// TIA Portal project "Plc_KTKDL" (V19) (continued)
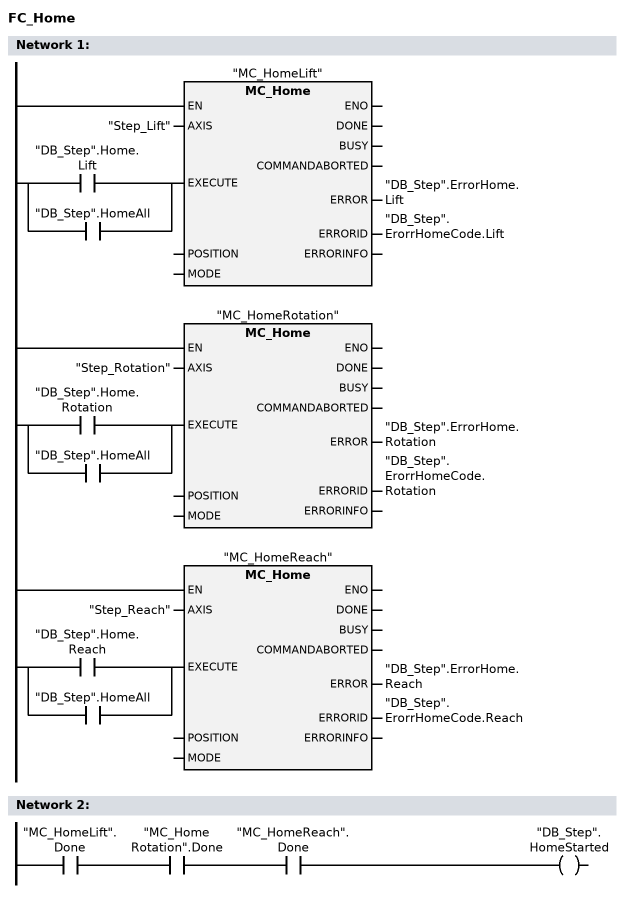
   "MC_HomeLift"(Axis := "Step_Lift",   // MC_Home
                 Execute := "DB_Step".Home.Lift OR "DB_Step".HomeAll,
                 Error => "DB_Step".ErrorHome.Lift,
                 ErrorID => "DB_Step".ErorrHomeCode.Lift);
   "MC_HomeRotation"(Axis := "Step_Rotation",   // MC_Home
                     Execute := "DB_Step".Home.Rotation OR "DB_Step".HomeAll,
                     Error => "DB_Step".ErrorHome.Rotation,
                     ErrorID => "DB_Step".ErorrHomeCode.Rotation);
   "MC_HomeReach"(Axis := "Step_Reach",   // MC_Home
                  Execute := "DB_Step".Home.Reach OR "DB_Step".HomeAll,
                  Error => "DB_Step".ErrorHome.Reach,
                  ErrorID => "DB_Step".ErorrHomeCode.Reach);
END_REGION

REGION Network 2
   RUNG wire#powerrail
      Contact( "MC_HomeLift".Done )
      Contact( "MC_HomeRotation".Done )
      Contact( "MC_HomeReach".Done )
      Coil( "DB_Step".HomeStarted )
   END_RUNG
   // the same network as SCL:
   "DB_Step".HomeStarted := "MC_HomeLift".Done AND "MC_HomeRotation".Done AND "MC_HomeReach".Done;
END_REGION
END_FUNCTION

FUNCTION "FC_Auto" : Void   // FC17, LAD
{ S7_Optimized_Access := 'TRUE' }
VERSION : 0.1
   VAR_TEMP   // added for the SCL form of the ladder/FBD networks
      _w1 : Bool;
      _w2 : Bool;
      _w3 : Bool;
      _w4 : Bool;
      _w5 : Bool;
      _w6 : Bool;
      _w7 : Bool;
      _w8 : Bool;
      _w9 : Bool;
      _w10 : Bool;
      _w11 : Bool;
      _w12 : Bool;
      _w13 : Bool;
      _w14 : Bool;
      _w15 : Bool;
      _w16 : Bool;
      _w17 : Bool;
      _w18 : Bool;
   END_VAR
BEGIN

REGION Network 1
   // 2 bước đầu là kiểm tra và set vận tốc
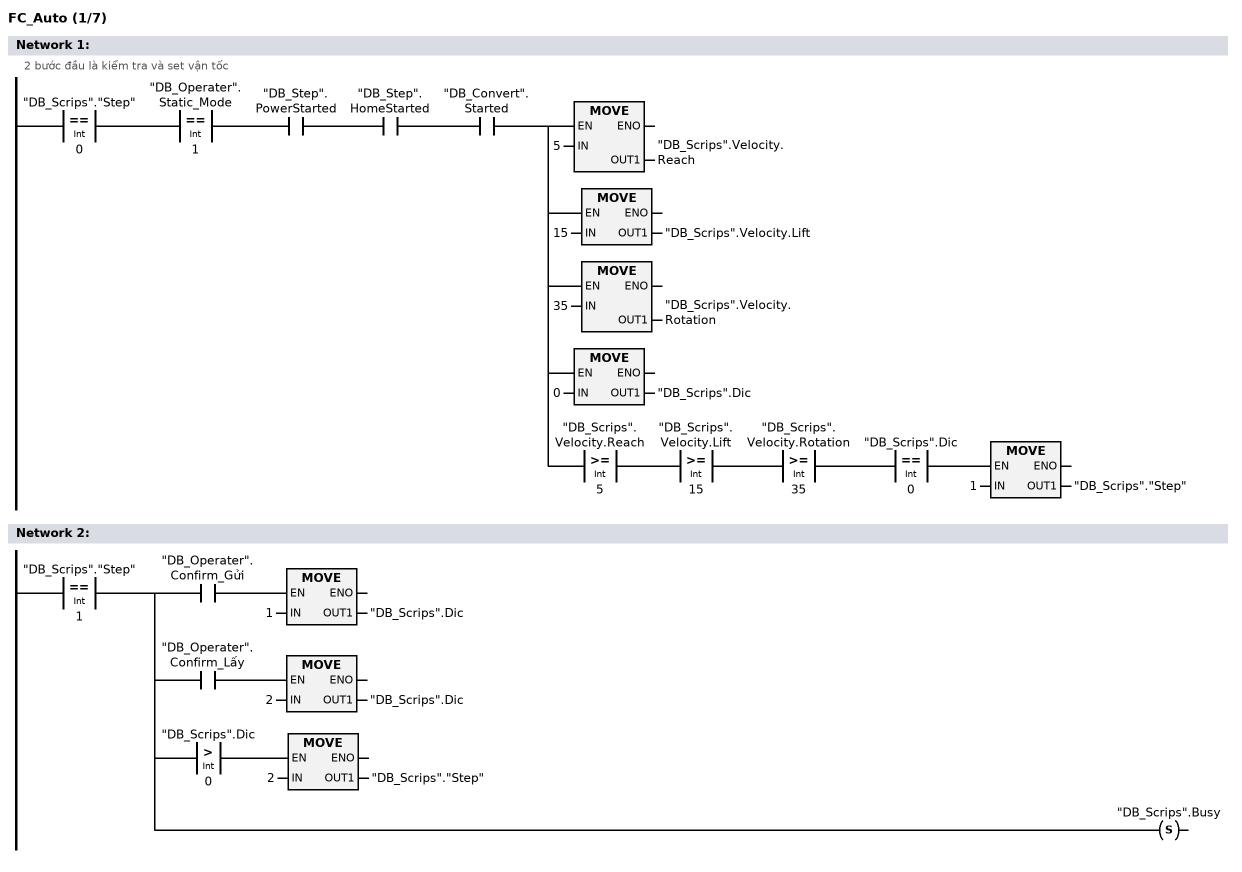
   RUNG wire#powerrail
      { S7_Templates := "SrcType := Int" } EQ_Contact(in1 := "DB_Scrips"."Step", in2 := 0)
      { S7_Templates := "SrcType := Int" } EQ_Contact(in1 := "DB_Operater".Static_Mode, in2 := 1)
      Contact( "DB_Step".PowerStarted )
      Contact( "DB_Step".HomeStarted )
      Contact( "DB_Convert".Started )
      wire#w1
      Move(in := 5, out1 => "DB_Scrips".Velocity.Reach)
   END_RUNG
   RUNG wire#w1
      Move(in := 15, out1 => "DB_Scrips".Velocity.Lift)
   END_RUNG
   RUNG wire#w1
      Move(in := 35, out1 => "DB_Scrips".Velocity.Rotation)
   END_RUNG
   RUNG wire#w1
      Move(in := 0, out1 => "DB_Scrips".Dic)
   END_RUNG
   RUNG wire#w1
      { S7_Templates := "SrcType := Int" } GE_Contact(in1 := "DB_Scrips".Velocity.Reach, in2 := 5)
      { S7_Templates := "SrcType := Int" } GE_Contact(in1 := "DB_Scrips".Velocity.Lift, in2 := 15)
      { S7_Templates := "SrcType := Int" } GE_Contact(in1 := "DB_Scrips".Velocity.Rotation, in2 := 35)
      { S7_Templates := "SrcType := Int" } EQ_Contact(in1 := "DB_Scrips".Dic, in2 := 0)
      Move(in := 1, out1 => "DB_Scrips"."Step")
   END_RUNG
   // the same network as SCL:
   #_w1 := ("DB_Scrips"."Step" = 0) AND ("DB_Operater".Static_Mode = 1) AND "DB_Step".PowerStarted AND "DB_Step".HomeStarted AND "DB_Convert".Started;
   IF #_w1 THEN
       "DB_Scrips".Velocity.Reach := 5;
       "DB_Scrips".Velocity.Lift := 15;
       "DB_Scrips".Velocity.Rotation := 35;
       "DB_Scrips".Dic := 0;
   END_IF;
   IF #_w1 AND ("DB_Scrips".Velocity.Reach >= 5) AND ("DB_Scrips".Velocity.Lift >= 15) AND ("DB_Scrips".Velocity.Rotation >= 35) AND ("DB_Scrips".Dic = 0) THEN
       "DB_Scrips"."Step" := 1;
   END_IF;
END_REGION

REGION Network 2
   RUNG wire#powerrail
      { S7_Templates := "SrcType := Int" } EQ_Contact(in1 := "DB_Scrips"."Step", in2 := 1)
      wire#w1
      Contact( "DB_Operater".Confirm_Gửi )
      Move(in := 1, out1 => "DB_Scrips".Dic)
   END_RUNG
   RUNG wire#w1
      Contact( "DB_Operater".Confirm_Lấy )
      Move(in := 2, out1 => "DB_Scrips".Dic)
   END_RUNG
   RUNG wire#w1
      { S7_Templates := "SrcType := Int" } GT_Contact(in1 := "DB_Scrips".Dic, in2 := 0)
      Move(in := 2, out1 => "DB_Scrips"."Step")
   END_RUNG
   RUNG wire#w1
      S_Coil( "DB_Scrips".Busy )
   END_RUNG
   // the same network as SCL:
   #_w1 := "DB_Scrips"."Step" = 1;
   IF #_w1 AND "DB_Operater".Confirm_Gửi THEN "DB_Scrips".Dic := 1; END_IF;
   IF #_w1 AND "DB_Operater".Confirm_Lấy THEN "DB_Scrips".Dic := 2; END_IF;
   IF #_w1 AND ("DB_Scrips".Dic > 0) THEN "DB_Scrips"."Step" := 2; END_IF;
   IF #_w1 THEN "DB_Scrips".Busy := TRUE; END_IF;
END_REGION

REGION Network 3
   // chưa làm logic lấy
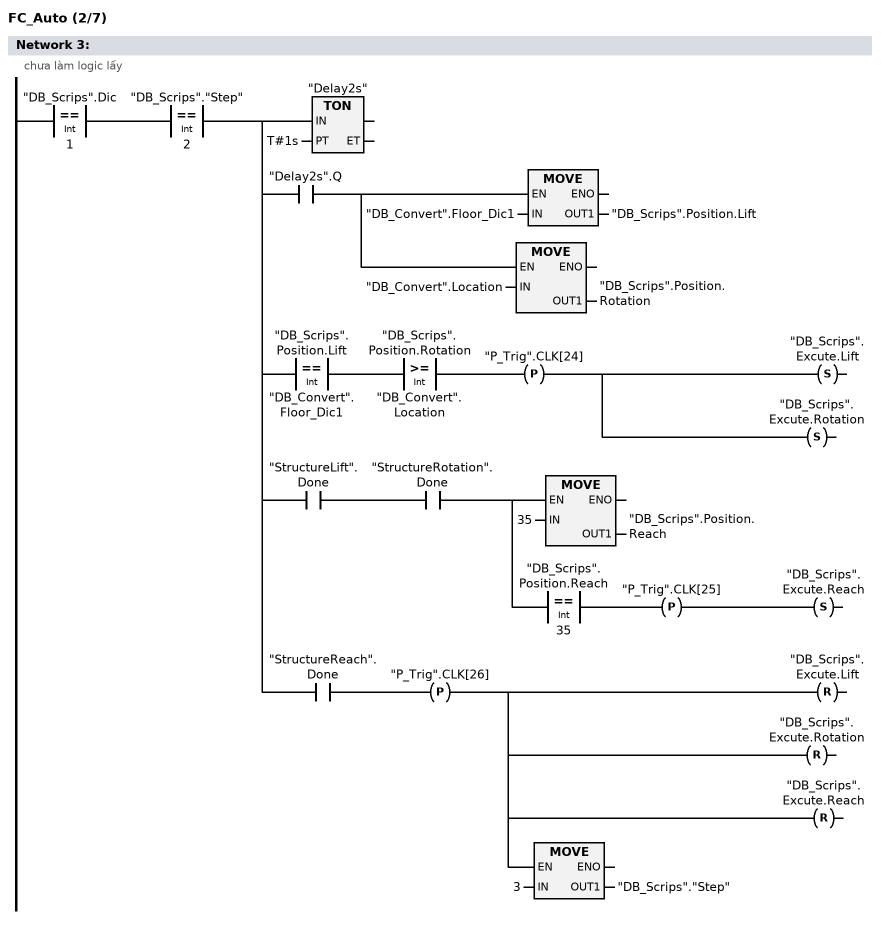
   #_w1 := ("DB_Scrips".Dic = 1) AND ("DB_Scrips"."Step" = 2);
   "Delay2s".TON(IN := #_w1, PT := T#1s);
   IF #_w1 AND "Delay2s".Q THEN
       "DB_Scrips".Position.Lift := "DB_Convert".Floor_Dic1;
       "DB_Scrips".Position.Rotation := "DB_Convert".Location;
   END_IF;
   #_w2 := #_w1 AND ("DB_Scrips".Position.Lift = "DB_Convert".Floor_Dic1) AND ("DB_Scrips".Position.Rotation >= "DB_Convert".Location);
   #_w3 := #_w2 AND NOT "P_Trig".CLK[24];   // rising edge
   "P_Trig".CLK[24] := #_w2;
   IF #_w3 THEN
       "DB_Scrips".Excute.Lift := TRUE;
       "DB_Scrips".Excute.Rotation := TRUE;
   END_IF;
   #_w4 := #_w1 AND "StructureLift".Done AND "StructureRotation".Done;
   IF #_w4 THEN "DB_Scrips".Position.Reach := 35; END_IF;
   #_w5 := #_w4 AND ("DB_Scrips".Position.Reach = 35);
   #_w6 := #_w5 AND NOT "P_Trig".CLK[25];   // rising edge
   "P_Trig".CLK[25] := #_w5;
   IF #_w6 THEN "DB_Scrips".Excute.Reach := TRUE; END_IF;
   #_w7 := #_w1 AND "StructureReach".Done;
   #_w8 := #_w7 AND NOT "P_Trig".CLK[26];   // rising edge
   "P_Trig".CLK[26] := #_w7;
   IF #_w8 THEN
       "DB_Scrips".Excute.Lift := FALSE;
       "DB_Scrips".Excute.Rotation := FALSE;
       "DB_Scrips".Excute.Reach := FALSE;
       "DB_Scrips"."Step" := 3;
   END_IF;
END_REGION

REGION Network 4
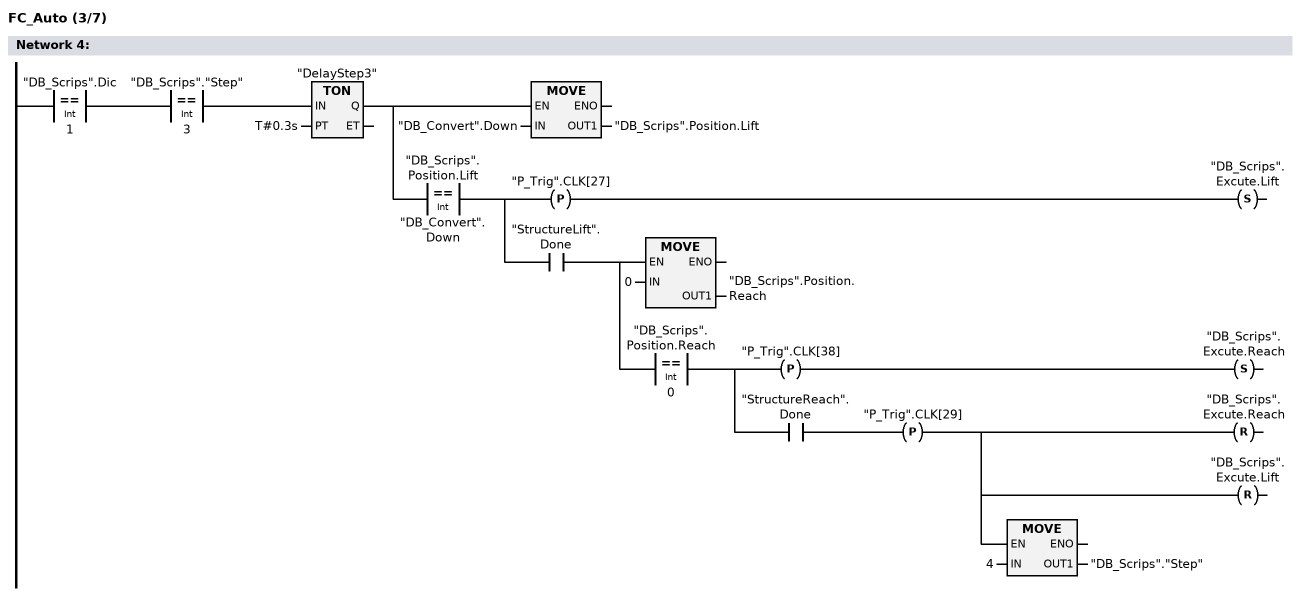
   "DelayStep3".TON(IN := ("DB_Scrips".Dic = 1) AND ("DB_Scrips"."Step" = 3), PT := T#0.3s);
   IF "DelayStep3".Q THEN "DB_Scrips".Position.Lift := "DB_Convert".Down; END_IF;
   #_w1 := "DelayStep3".Q AND ("DB_Scrips".Position.Lift = "DB_Convert".Down);
   #_w2 := #_w1 AND NOT "P_Trig".CLK[27];   // rising edge
   "P_Trig".CLK[27] := #_w1;
   IF #_w2 THEN "DB_Scrips".Excute.Lift := TRUE; END_IF;
   #_w3 := #_w1 AND "StructureLift".Done;
   IF #_w3 THEN "DB_Scrips".Position.Reach := 0; END_IF;
   #_w4 := #_w3 AND ("DB_Scrips".Position.Reach = 0);
   #_w5 := #_w4 AND NOT "P_Trig".CLK[38];   // rising edge
   "P_Trig".CLK[38] := #_w4;
   IF #_w5 THEN "DB_Scrips".Excute.Reach := TRUE; END_IF;
   #_w6 := #_w4 AND "StructureReach".Done;
   #_w7 := #_w6 AND NOT "P_Trig".CLK[29];   // rising edge
   "P_Trig".CLK[29] := #_w6;
   IF #_w7 THEN
       "DB_Scrips".Excute.Reach := FALSE;
       "DB_Scrips".Excute.Lift := FALSE;
       "DB_Scrips"."Step" := 4;
   END_IF;
END_REGION

REGION Network 5
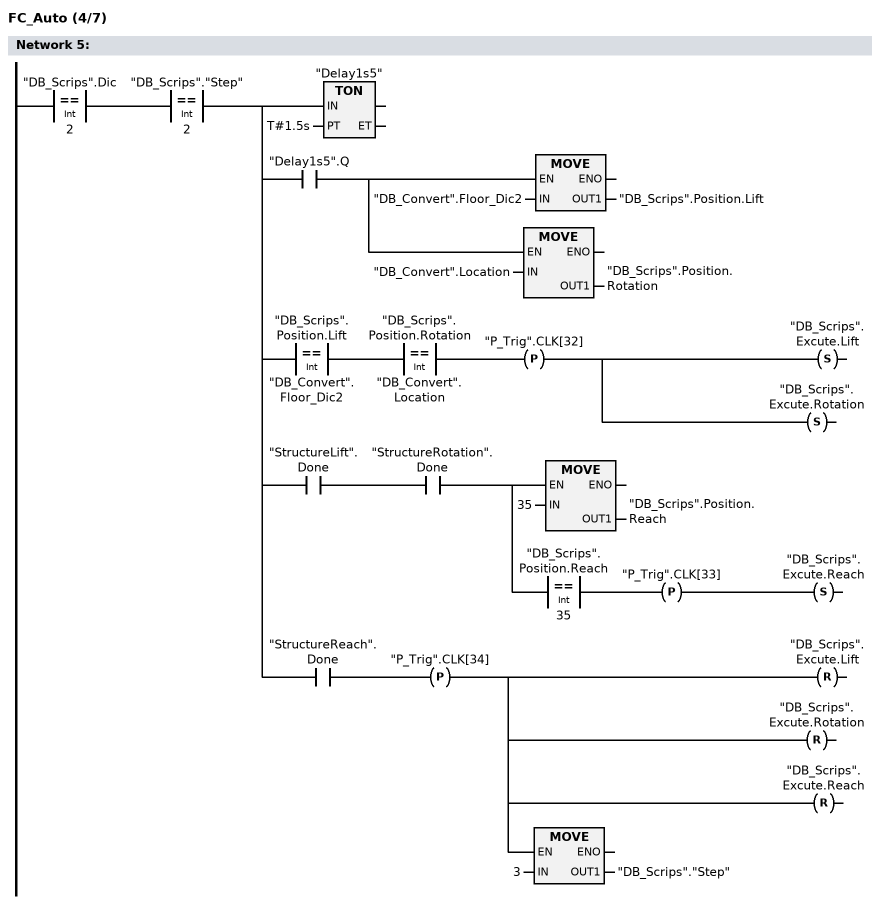
   #_w1 := ("DB_Scrips".Dic = 2) AND ("DB_Scrips"."Step" = 2);
   "Delay1s5".TON(IN := #_w1, PT := T#1.5s);
   IF #_w1 AND "Delay1s5".Q THEN
       "DB_Scrips".Position.Lift := "DB_Convert".Floor_Dic2;
       "DB_Scrips".Position.Rotation := "DB_Convert".Location;
   END_IF;
   #_w2 := #_w1 AND ("DB_Scrips".Position.Lift = "DB_Convert".Floor_Dic2) AND ("DB_Scrips".Position.Rotation = "DB_Convert".Location);
   #_w3 := #_w2 AND NOT "P_Trig".CLK[32];   // rising edge
   "P_Trig".CLK[32] := #_w2;
   IF #_w3 THEN
       "DB_Scrips".Excute.Lift := TRUE;
       "DB_Scrips".Excute.Rotation := TRUE;
   END_IF;
   #_w4 := #_w1 AND "StructureLift".Done AND "StructureRotation".Done;
   IF #_w4 THEN "DB_Scrips".Position.Reach := 35; END_IF;
   #_w5 := #_w4 AND ("DB_Scrips".Position.Reach = 35);
   #_w6 := #_w5 AND NOT "P_Trig".CLK[33];   // rising edge
   "P_Trig".CLK[33] := #_w5;
   IF #_w6 THEN "DB_Scrips".Excute.Reach := TRUE; END_IF;
   #_w7 := #_w1 AND "StructureReach".Done;
   #_w8 := #_w7 AND NOT "P_Trig".CLK[34];   // rising edge
   "P_Trig".CLK[34] := #_w7;
   IF #_w8 THEN
       "DB_Scrips".Excute.Lift := FALSE;
       "DB_Scrips".Excute.Rotation := FALSE;
       "DB_Scrips".Excute.Reach := FALSE;
       "DB_Scrips"."Step" := 3;
   END_IF;
END_REGION

REGION Network 6
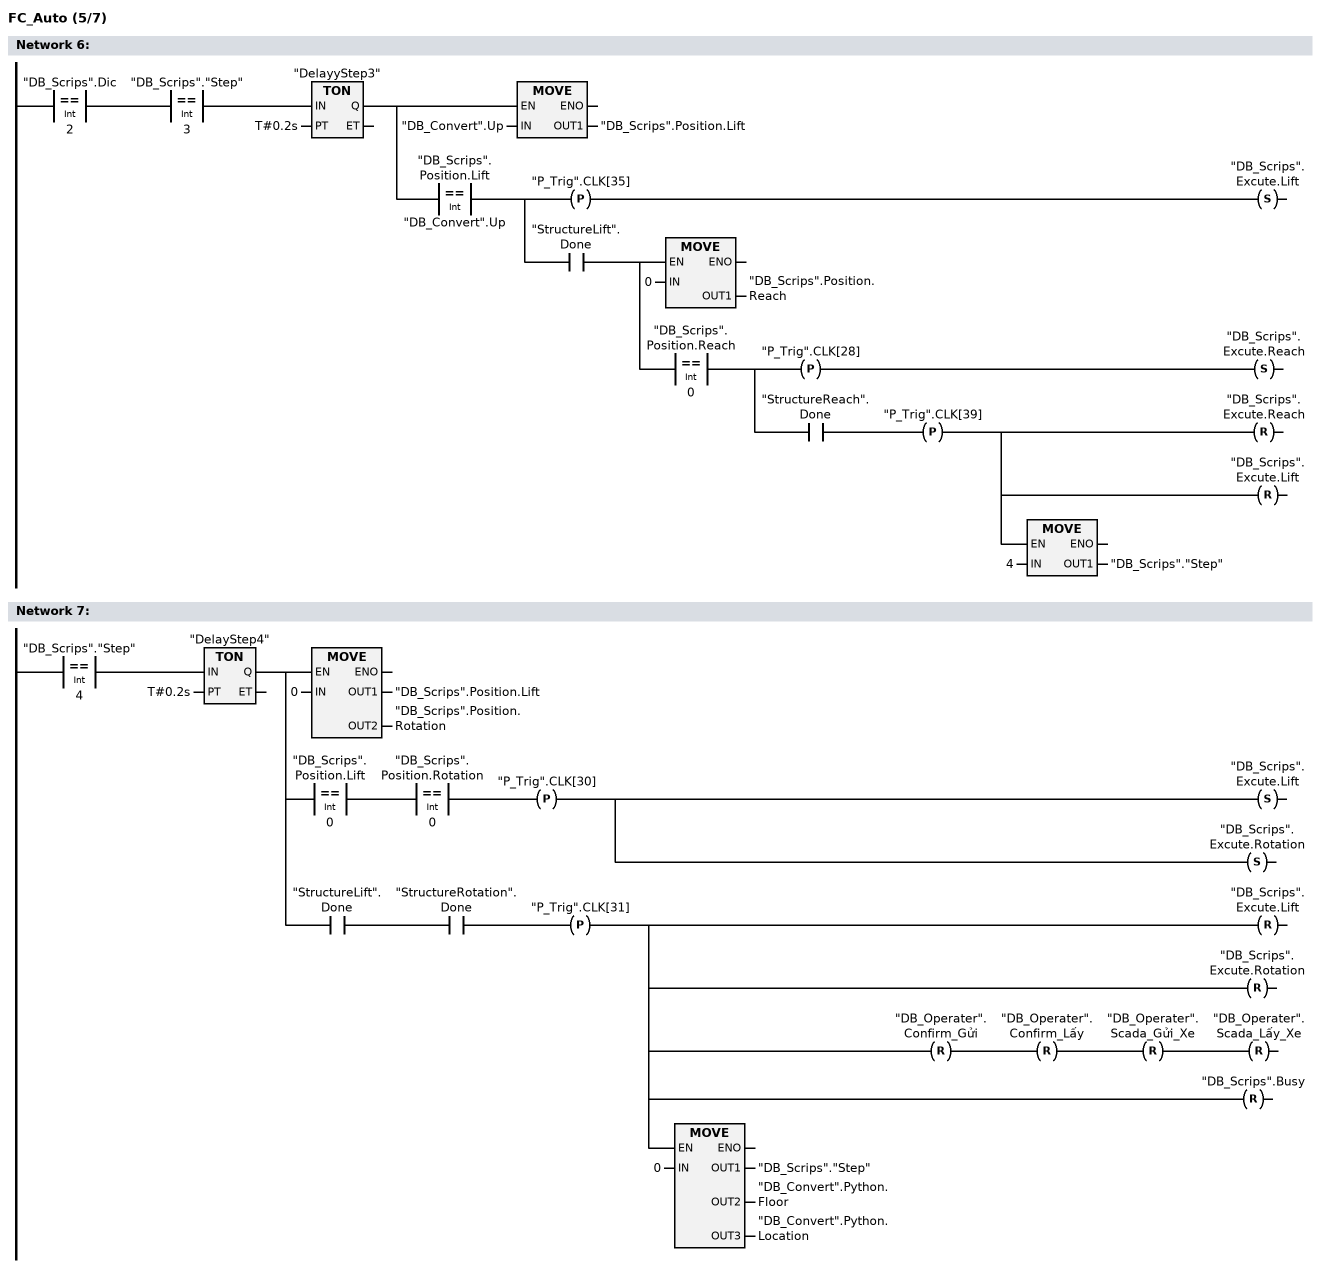
   "DelayyStep3".TON(IN := ("DB_Scrips".Dic = 2) AND ("DB_Scrips"."Step" = 3), PT := T#0.2s);
   IF "DelayyStep3".Q THEN "DB_Scrips".Position.Lift := "DB_Convert".Up; END_IF;
   #_w1 := "DelayyStep3".Q AND ("DB_Scrips".Position.Lift = "DB_Convert".Up);
   #_w2 := #_w1 AND NOT "P_Trig".CLK[35];   // rising edge
   "P_Trig".CLK[35] := #_w1;
   IF #_w2 THEN "DB_Scrips".Excute.Lift := TRUE; END_IF;
   #_w3 := #_w1 AND "StructureLift".Done;
   IF #_w3 THEN "DB_Scrips".Position.Reach := 0; END_IF;
   #_w4 := #_w3 AND ("DB_Scrips".Position.Reach = 0);
   #_w5 := #_w4 AND NOT "P_Trig".CLK[28];   // rising edge
   "P_Trig".CLK[28] := #_w4;
   IF #_w5 THEN "DB_Scrips".Excute.Reach := TRUE; END_IF;
   #_w6 := #_w4 AND "StructureReach".Done;
   #_w7 := #_w6 AND NOT "P_Trig".CLK[39];   // rising edge
   "P_Trig".CLK[39] := #_w6;
   IF #_w7 THEN
       "DB_Scrips".Excute.Reach := FALSE;
       "DB_Scrips".Excute.Lift := FALSE;
       "DB_Scrips"."Step" := 4;
   END_IF;
END_REGION

REGION Network 7
   "DelayStep4".TON(IN := "DB_Scrips"."Step" = 4, PT := T#0.2s);
   IF "DelayStep4".Q THEN
       "DB_Scrips".Position.Lift := 0;
       "DB_Scrips".Position.Rotation := 0;
   END_IF;
   #_w1 := "DelayStep4".Q AND ("DB_Scrips".Position.Lift = 0) AND ("DB_Scrips".Position.Rotation = 0);
   #_w2 := #_w1 AND NOT "P_Trig".CLK[30];   // rising edge
   "P_Trig".CLK[30] := #_w1;
   IF #_w2 THEN
       "DB_Scrips".Excute.Lift := TRUE;
       "DB_Scrips".Excute.Rotation := TRUE;
   END_IF;
   #_w3 := "DelayStep4".Q AND "StructureLift".Done AND "StructureRotation".Done;
   #_w4 := #_w3 AND NOT "P_Trig".CLK[31];   // rising edge
   "P_Trig".CLK[31] := #_w3;
   IF #_w4 THEN
       "DB_Scrips".Excute.Lift := FALSE;
       "DB_Scrips".Excute.Rotation := FALSE;
       "DB_Operater".Confirm_Gửi := FALSE;
       "DB_Operater".Confirm_Lấy := FALSE;
       "DB_Operater".Scada_Gửi_Xe := FALSE;
       "DB_Operater".Scada_Lấy_Xe := FALSE;
       "DB_Scrips".Busy := FALSE;
       "DB_Scrips"."Step" := 0;
       "DB_Convert".Python.Floor := 0;
       "DB_Convert".Python.Location := 0;
   END_IF;
END_REGION

REGION Network 9
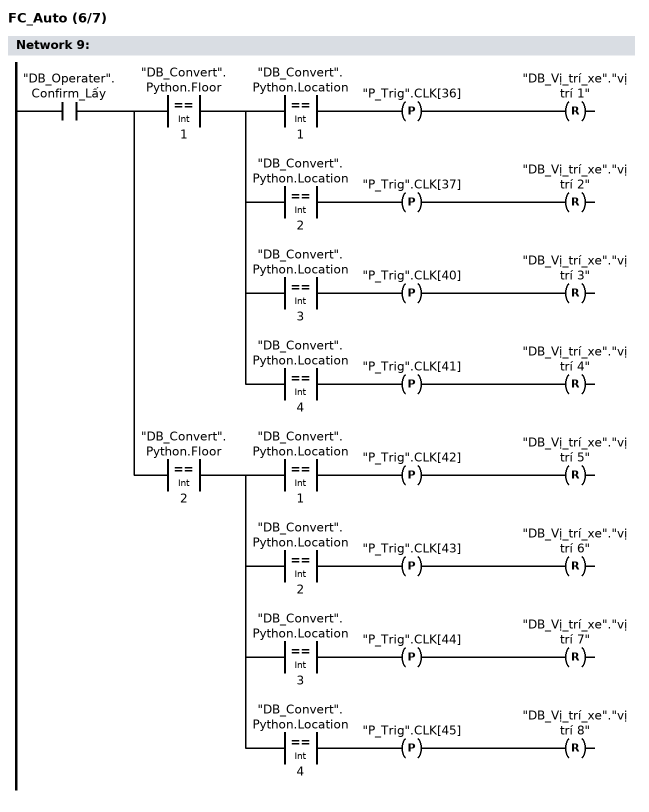
   RUNG wire#powerrail
      Contact( "DB_Operater".Confirm_Lấy )
      wire#w1
      { S7_Templates := "SrcType := Int" } EQ_Contact(in1 := "DB_Convert".Python.Floor, in2 := 1)
      wire#w2
      { S7_Templates := "SrcType := Int" } EQ_Contact(in1 := "DB_Convert".Python.Location, in2 := 1)
      P_Trig( "P_Trig".CLK[36] )
      R_Coil( "DB_Vị_trí_xe"."vị trí 1" )
   END_RUNG
   RUNG wire#w2
      { S7_Templates := "SrcType := Int" } EQ_Contact(in1 := "DB_Convert".Python.Location, in2 := 2)
      P_Trig( "P_Trig".CLK[37] )
      R_Coil( "DB_Vị_trí_xe"."vị trí 2" )
   END_RUNG
   RUNG wire#w2
      { S7_Templates := "SrcType := Int" } EQ_Contact(in1 := "DB_Convert".Python.Location, in2 := 3)
      P_Trig( "P_Trig".CLK[40] )
      R_Coil( "DB_Vị_trí_xe"."vị trí 3" )
   END_RUNG
   RUNG wire#w2
      { S7_Templates := "SrcType := Int" } EQ_Contact(in1 := "DB_Convert".Python.Location, in2 := 4)
      P_Trig( "P_Trig".CLK[41] )
      R_Coil( "DB_Vị_trí_xe"."vị trí 4" )
   END_RUNG
   RUNG wire#w1
      { S7_Templates := "SrcType := Int" } EQ_Contact(in1 := "DB_Convert".Python.Floor, in2 := 2)
      wire#w3
      { S7_Templates := "SrcType := Int" } EQ_Contact(in1 := "DB_Convert".Python.Location, in2 := 1)
      P_Trig( "P_Trig".CLK[42] )
      R_Coil( "DB_Vị_trí_xe"."vị trí 5" )
   END_RUNG
   RUNG wire#w3
      { S7_Templates := "SrcType := Int" } EQ_Contact(in1 := "DB_Convert".Python.Location, in2 := 2)
      P_Trig( "P_Trig".CLK[43] )
      R_Coil( "DB_Vị_trí_xe"."vị trí 6" )
   END_RUNG
   RUNG wire#w3
      { S7_Templates := "SrcType := Int" } EQ_Contact(in1 := "DB_Convert".Python.Location, in2 := 3)
      P_Trig( "P_Trig".CLK[44] )
      R_Coil( "DB_Vị_trí_xe"."vị trí 7" )
   END_RUNG
   RUNG wire#w3
      { S7_Templates := "SrcType := Int" } EQ_Contact(in1 := "DB_Convert".Python.Location, in2 := 4)
      P_Trig( "P_Trig".CLK[45] )
      R_Coil( "DB_Vị_trí_xe"."vị trí 8" )
   END_RUNG
   // the same network as SCL:
   #_w1 := "DB_Operater".Confirm_Lấy AND ("DB_Convert".Python.Floor = 1);
   #_w2 := #_w1 AND ("DB_Convert".Python.Location = 1);
   #_w3 := #_w2 AND NOT "P_Trig".CLK[36];   // rising edge
   "P_Trig".CLK[36] := #_w2;
   IF #_w3 THEN "DB_Vị_trí_xe"."vị trí 1" := FALSE; END_IF;
   #_w4 := #_w1 AND ("DB_Convert".Python.Location = 2);
   #_w5 := #_w4 AND NOT "P_Trig".CLK[37];   // rising edge
   "P_Trig".CLK[37] := #_w4;
   IF #_w5 THEN "DB_Vị_trí_xe"."vị trí 2" := FALSE; END_IF;
   #_w6 := #_w1 AND ("DB_Convert".Python.Location = 3);
   #_w7 := #_w6 AND NOT "P_Trig".CLK[40];   // rising edge
   "P_Trig".CLK[40] := #_w6;
   IF #_w7 THEN "DB_Vị_trí_xe"."vị trí 3" := FALSE; END_IF;
   #_w8 := #_w1 AND ("DB_Convert".Python.Location = 4);
   #_w9 := #_w8 AND NOT "P_Trig".CLK[41];   // rising edge
   "P_Trig".CLK[41] := #_w8;
   IF #_w9 THEN "DB_Vị_trí_xe"."vị trí 4" := FALSE; END_IF;
   #_w10 := "DB_Operater".Confirm_Lấy AND ("DB_Convert".Python.Floor = 2);
   #_w11 := #_w10 AND ("DB_Convert".Python.Location = 1);
   #_w12 := #_w11 AND NOT "P_Trig".CLK[42];   // rising edge
   "P_Trig".CLK[42] := #_w11;
   IF #_w12 THEN "DB_Vị_trí_xe"."vị trí 5" := FALSE; END_IF;
   #_w13 := #_w10 AND ("DB_Convert".Python.Location = 2);
   #_w14 := #_w13 AND NOT "P_Trig".CLK[43];   // rising edge
   "P_Trig".CLK[43] := #_w13;
   IF #_w14 THEN "DB_Vị_trí_xe"."vị trí 6" := FALSE; END_IF;
   #_w15 := #_w10 AND ("DB_Convert".Python.Location = 3);
   #_w16 := #_w15 AND NOT "P_Trig".CLK[44];   // rising edge
   "P_Trig".CLK[44] := #_w15;
   IF #_w16 THEN "DB_Vị_trí_xe"."vị trí 7" := FALSE; END_IF;
   #_w17 := #_w10 AND ("DB_Convert".Python.Location = 4);
   #_w18 := #_w17 AND NOT "P_Trig".CLK[45];   // rising edge
   "P_Trig".CLK[45] := #_w17;
   IF #_w18 THEN "DB_Vị_trí_xe"."vị trí 8" := FALSE; END_IF;
END_REGION

REGION Network 10
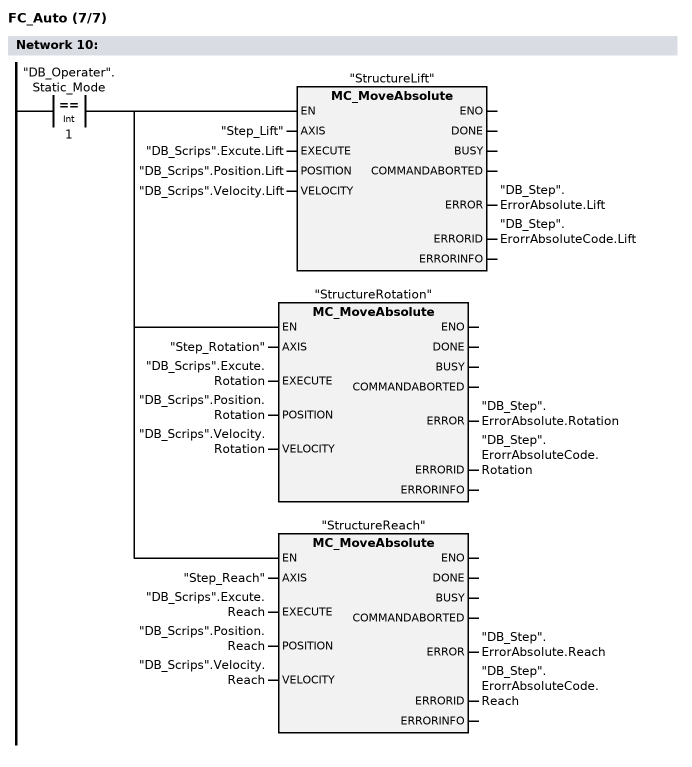
   #_w1 := "DB_Operater".Static_Mode = 1;
   IF #_w1 THEN
       "StructureLift"(Axis := "Step_Lift",   // MC_MoveAbsolute
                       Execute := "DB_Scrips".Excute.Lift,
                       Position := "DB_Scrips".Position.Lift,
                       Velocity := "DB_Scrips".Velocity.Lift,
                       Error => "DB_Step".ErrorAbsolute.Lift,
                       ErrorID => "DB_Step".ErorrAbsoluteCode.Lift);
       "StructureRotation"(Axis := "Step_Rotation",   // MC_MoveAbsolute
                           Execute := "DB_Scrips".Excute.Rotation,
                           Position := "DB_Scrips".Position.Rotation,
                           Velocity := "DB_Scrips".Velocity.Rotation,
                           Error => "DB_Step".ErrorAbsolute.Rotation,
                           ErrorID => "DB_Step".ErorrAbsoluteCode.Rotation);
       "StructureReach"(Axis := "Step_Reach",   // MC_MoveAbsolute
                        Execute := "DB_Scrips".Excute.Reach,
                        Position := "DB_Scrips".Position.Reach,
                        Velocity := "DB_Scrips".Velocity.Reach,
                        Error => "DB_Step".ErrorAbsolute.Reach,
                        ErrorID => "DB_Step".ErorrAbsoluteCode.Reach);
   END_IF;
END_REGION
END_FUNCTION

FUNCTION "FC_Reset" : Void   // FC18, LAD
{ S7_Optimized_Access := 'TRUE' }
VERSION : 0.1
BEGIN

REGION Network 1
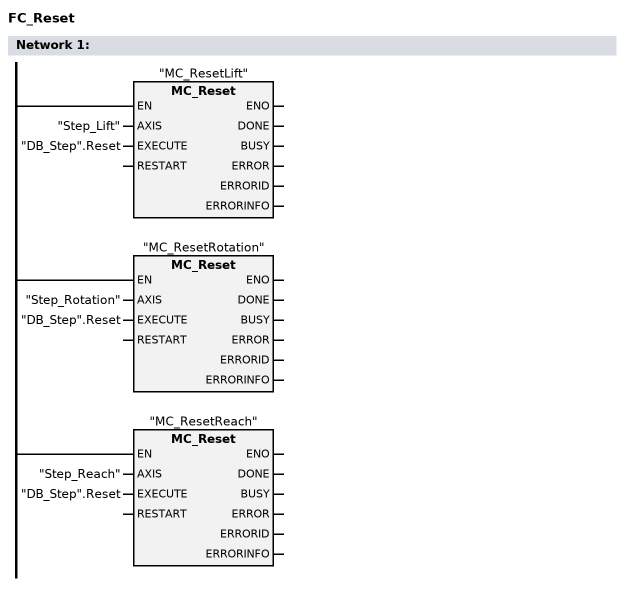
   "MC_ResetLift"(Axis := "Step_Lift", Execute := "DB_Step".Reset);   // MC_Reset
   "MC_ResetRotation"(Axis := "Step_Rotation", Execute := "DB_Step".Reset);   // MC_Reset
   "MC_ResetReach"(Axis := "Step_Reach", Execute := "DB_Step".Reset);   // MC_Reset
END_REGION
END_FUNCTION

// folder: đầy , các logic tìm

FUNCTION "FC_Tìm_tầng" : Void   // FC2, LAD
{ S7_Optimized_Access := 'TRUE' }
VERSION : 0.1
   VAR_TEMP   // added for the SCL form of the ladder/FBD networks
      _w1 : Bool;
      _w2 : Bool;
      _w3 : Bool;
      _w4 : Bool;
      _w5 : Bool;
   END_VAR
BEGIN

REGION Network 1
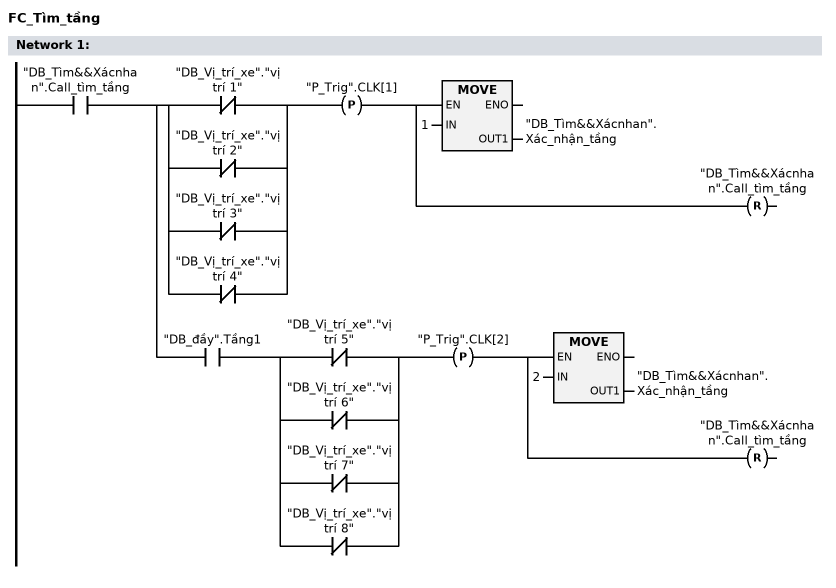
   RUNG wire#powerrail
      Contact( "DB_Tìm&&Xácnhan".Call_tìm_tầng )
      wire#w1
      I_Contact( "DB_Vị_trí_xe"."vị trí 1" )
      wire#w2
      P_Trig( "P_Trig".CLK[1] )
      wire#w3
      Move(in := 1, out1 => "DB_Tìm&&Xácnhan".Xác_nhận_tầng)
   END_RUNG
   RUNG wire#w1
      I_Contact( "DB_Vị_trí_xe"."vị trí 2" )
   END_RUNG wire#w2
   RUNG wire#w1
      I_Contact( "DB_Vị_trí_xe"."vị trí 3" )
   END_RUNG wire#w2
   RUNG wire#w1
      I_Contact( "DB_Vị_trí_xe"."vị trí 4" )
   END_RUNG wire#w2
   RUNG wire#w3
      R_Coil( "DB_Tìm&&Xácnhan".Call_tìm_tầng )
   END_RUNG
   RUNG wire#w1
      Contact( "DB_đầy".Tầng1 )
      wire#w4
      I_Contact( "DB_Vị_trí_xe"."vị trí 5" )
      wire#w5
      P_Trig( "P_Trig".CLK[2] )
      wire#w6
      Move(in := 2, out1 => "DB_Tìm&&Xácnhan".Xác_nhận_tầng)
   END_RUNG
   RUNG wire#w4
      I_Contact( "DB_Vị_trí_xe"."vị trí 6" )
   END_RUNG wire#w5
   RUNG wire#w4
      I_Contact( "DB_Vị_trí_xe"."vị trí 7" )
   END_RUNG wire#w5
   RUNG wire#w4
      I_Contact( "DB_Vị_trí_xe"."vị trí 8" )
   END_RUNG wire#w5
   RUNG wire#w6
      R_Coil( "DB_Tìm&&Xácnhan".Call_tìm_tầng )
   END_RUNG
   // the same network as SCL:
   #_w1 := "DB_Tìm&&Xácnhan".Call_tìm_tầng AND (NOT "DB_Vị_trí_xe"."vị trí 1" OR NOT "DB_Vị_trí_xe"."vị trí 2" OR NOT "DB_Vị_trí_xe"."vị trí 3" OR NOT "DB_Vị_trí_xe"."vị trí 4");
   #_w2 := #_w1 AND NOT "P_Trig".CLK[1];   // rising edge
   "P_Trig".CLK[1] := #_w1;
   IF #_w2 THEN "DB_Tìm&&Xácnhan".Xác_nhận_tầng := 1; END_IF;
   #_w3 := "DB_Tìm&&Xácnhan".Call_tìm_tầng;
   IF #_w2 THEN "DB_Tìm&&Xácnhan".Call_tìm_tầng := FALSE; END_IF;
   #_w4 := #_w3 AND "DB_đầy".Tầng1 AND (NOT "DB_Vị_trí_xe"."vị trí 5" OR NOT "DB_Vị_trí_xe"."vị trí 6" OR NOT "DB_Vị_trí_xe"."vị trí 7" OR NOT "DB_Vị_trí_xe"."vị trí 8");
   #_w5 := #_w4 AND NOT "P_Trig".CLK[2];   // rising edge
   "P_Trig".CLK[2] := #_w4;
   IF #_w5 THEN
       "DB_Tìm&&Xácnhan".Xác_nhận_tầng := 2;
       "DB_Tìm&&Xácnhan".Call_tìm_tầng := FALSE;
   END_IF;
END_REGION
END_FUNCTION

FUNCTION "FC_Tìm_vị_trí_tầng1" : Void   // FC3, LAD
{ S7_Optimized_Access := 'TRUE' }
VERSION : 0.1
   VAR_TEMP   // added for the SCL form of the ladder/FBD networks
      _w1 : Bool;
      _w2 : Bool;
   END_VAR
BEGIN

REGION Network 1
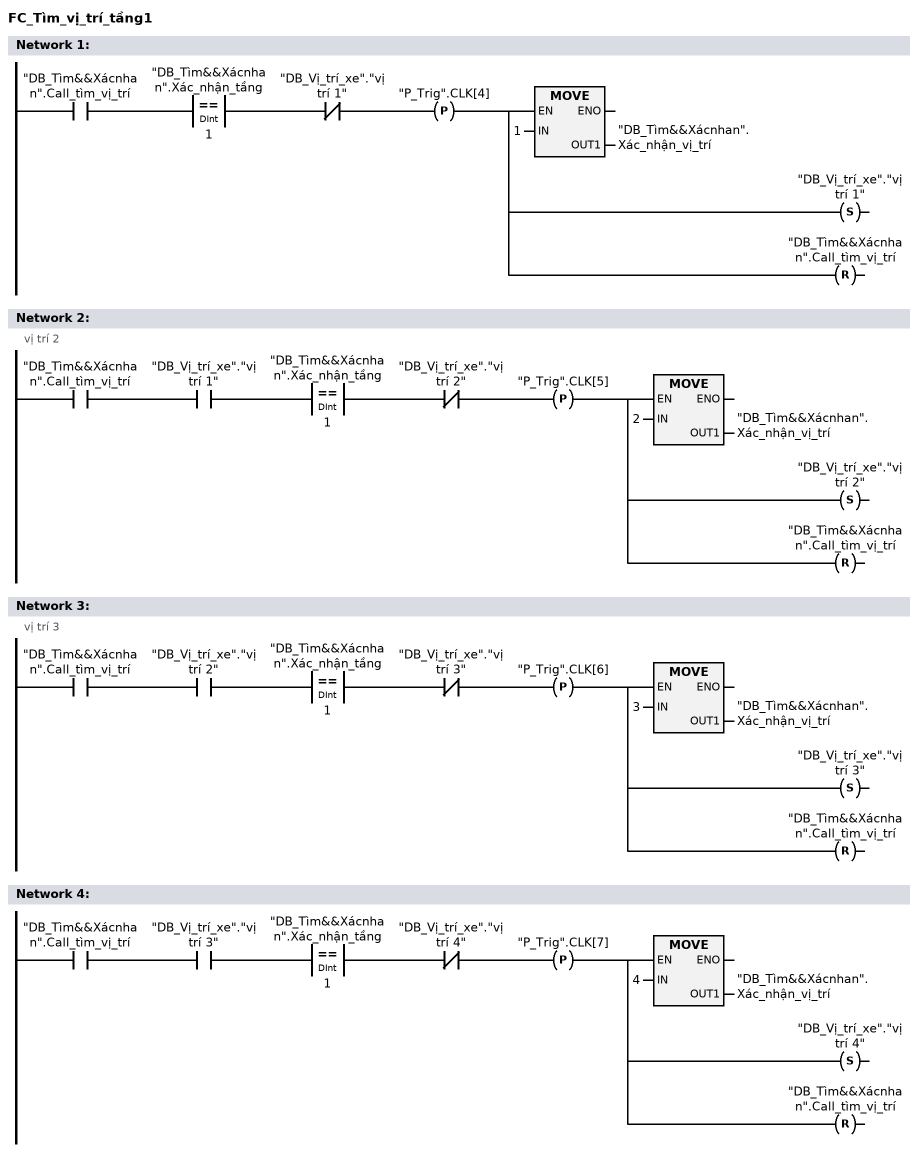
   RUNG wire#powerrail
      Contact( "DB_Tìm&&Xácnhan".Call_tìm_vị_trí )
      { S7_Templates := "SrcType := DInt" } EQ_Contact(in1 := "DB_Tìm&&Xácnhan".Xác_nhận_tầng, in2 := 1)
      I_Contact( "DB_Vị_trí_xe"."vị trí 1" )
      P_Trig( "P_Trig".CLK[4] )
      wire#w1
      Move(in := 1, out1 => "DB_Tìm&&Xácnhan".Xác_nhận_vị_trí)
   END_RUNG
   RUNG wire#w1
      S_Coil( "DB_Vị_trí_xe"."vị trí 1" )
   END_RUNG
   RUNG wire#w1
      R_Coil( "DB_Tìm&&Xácnhan".Call_tìm_vị_trí )
   END_RUNG
   // the same network as SCL:
   #_w1 := "DB_Tìm&&Xácnhan".Call_tìm_vị_trí AND ("DB_Tìm&&Xácnhan".Xác_nhận_tầng = 1) AND NOT "DB_Vị_trí_xe"."vị trí 1";
   #_w2 := #_w1 AND NOT "P_Trig".CLK[4];   // rising edge
   "P_Trig".CLK[4] := #_w1;
   IF #_w2 THEN
       "DB_Tìm&&Xácnhan".Xác_nhận_vị_trí := 1;
       "DB_Vị_trí_xe"."vị trí 1" := TRUE;
       "DB_Tìm&&Xácnhan".Call_tìm_vị_trí := FALSE;
   END_IF;
END_REGION

REGION Network 2
   // vị trí 2
   RUNG wire#powerrail
      Contact( "DB_Tìm&&Xácnhan".Call_tìm_vị_trí )
      Contact( "DB_Vị_trí_xe"."vị trí 1" )
      { S7_Templates := "SrcType := DInt" } EQ_Contact(in1 := "DB_Tìm&&Xácnhan".Xác_nhận_tầng, in2 := 1)
      I_Contact( "DB_Vị_trí_xe"."vị trí 2" )
      P_Trig( "P_Trig".CLK[5] )
      wire#w1
      Move(in := 2, out1 => "DB_Tìm&&Xácnhan".Xác_nhận_vị_trí)
   END_RUNG
   RUNG wire#w1
      S_Coil( "DB_Vị_trí_xe"."vị trí 2" )
   END_RUNG
   RUNG wire#w1
      R_Coil( "DB_Tìm&&Xácnhan".Call_tìm_vị_trí )
   END_RUNG
   // the same network as SCL:
   #_w1 := "DB_Tìm&&Xácnhan".Call_tìm_vị_trí AND "DB_Vị_trí_xe"."vị trí 1" AND ("DB_Tìm&&Xácnhan".Xác_nhận_tầng = 1) AND NOT "DB_Vị_trí_xe"."vị trí 2";
   #_w2 := #_w1 AND NOT "P_Trig".CLK[5];   // rising edge
   "P_Trig".CLK[5] := #_w1;
   IF #_w2 THEN
       "DB_Tìm&&Xácnhan".Xác_nhận_vị_trí := 2;
       "DB_Vị_trí_xe"."vị trí 2" := TRUE;
       "DB_Tìm&&Xácnhan".Call_tìm_vị_trí := FALSE;
   END_IF;
END_REGION

REGION Network 3
   // vị trí 3
   RUNG wire#powerrail
      Contact( "DB_Tìm&&Xácnhan".Call_tìm_vị_trí )
      Contact( "DB_Vị_trí_xe"."vị trí 2" )
      { S7_Templates := "SrcType := DInt" } EQ_Contact(in1 := "DB_Tìm&&Xácnhan".Xác_nhận_tầng, in2 := 1)
      I_Contact( "DB_Vị_trí_xe"."vị trí 3" )
      P_Trig( "P_Trig".CLK[6] )
      wire#w1
      Move(in := 3, out1 => "DB_Tìm&&Xácnhan".Xác_nhận_vị_trí)
   END_RUNG
   RUNG wire#w1
      S_Coil( "DB_Vị_trí_xe"."vị trí 3" )
   END_RUNG
   RUNG wire#w1
      R_Coil( "DB_Tìm&&Xácnhan".Call_tìm_vị_trí )
   END_RUNG
   // the same network as SCL:
   #_w1 := "DB_Tìm&&Xácnhan".Call_tìm_vị_trí AND "DB_Vị_trí_xe"."vị trí 2" AND ("DB_Tìm&&Xácnhan".Xác_nhận_tầng = 1) AND NOT "DB_Vị_trí_xe"."vị trí 3";
   #_w2 := #_w1 AND NOT "P_Trig".CLK[6];   // rising edge
   "P_Trig".CLK[6] := #_w1;
   IF #_w2 THEN
       "DB_Tìm&&Xácnhan".Xác_nhận_vị_trí := 3;
       "DB_Vị_trí_xe"."vị trí 3" := TRUE;
       "DB_Tìm&&Xácnhan".Call_tìm_vị_trí := FALSE;
   END_IF;
END_REGION

REGION Network 4
   RUNG wire#powerrail
      Contact( "DB_Tìm&&Xácnhan".Call_tìm_vị_trí )
      Contact( "DB_Vị_trí_xe"."vị trí 3" )
      { S7_Templates := "SrcType := DInt" } EQ_Contact(in1 := "DB_Tìm&&Xácnhan".Xác_nhận_tầng, in2 := 1)
      I_Contact( "DB_Vị_trí_xe"."vị trí 4" )
      P_Trig( "P_Trig".CLK[7] )
      wire#w1
      Move(in := 4, out1 => "DB_Tìm&&Xácnhan".Xác_nhận_vị_trí)
   END_RUNG
   RUNG wire#w1
      S_Coil( "DB_Vị_trí_xe"."vị trí 4" )
   END_RUNG
   RUNG wire#w1
      R_Coil( "DB_Tìm&&Xácnhan".Call_tìm_vị_trí )
   END_RUNG
   // the same network as SCL:
   #_w1 := "DB_Tìm&&Xácnhan".Call_tìm_vị_trí AND "DB_Vị_trí_xe"."vị trí 3" AND ("DB_Tìm&&Xácnhan".Xác_nhận_tầng = 1) AND NOT "DB_Vị_trí_xe"."vị trí 4";
   #_w2 := #_w1 AND NOT "P_Trig".CLK[7];   // rising edge
   "P_Trig".CLK[7] := #_w1;
   IF #_w2 THEN
       "DB_Tìm&&Xácnhan".Xác_nhận_vị_trí := 4;
       "DB_Vị_trí_xe"."vị trí 4" := TRUE;
       "DB_Tìm&&Xácnhan".Call_tìm_vị_trí := FALSE;
   END_IF;
END_REGION
END_FUNCTION

FUNCTION "FC_đầy" : Void   // FC4, LAD
{ S7_Optimized_Access := 'TRUE' }
VERSION : 0.1
BEGIN

REGION Network 1
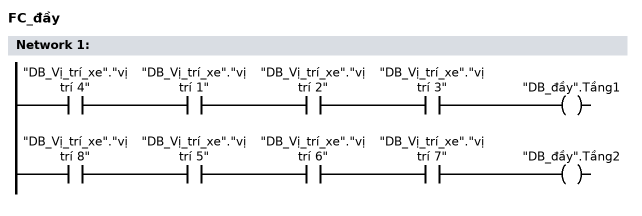
   RUNG wire#powerrail
      Contact( "DB_Vị_trí_xe"."vị trí 4" )
      Contact( "DB_Vị_trí_xe"."vị trí 1" )
      Contact( "DB_Vị_trí_xe"."vị trí 2" )
      Contact( "DB_Vị_trí_xe"."vị trí 3" )
      Coil( "DB_đầy".Tầng1 )
   END_RUNG
   RUNG wire#powerrail
      Contact( "DB_Vị_trí_xe"."vị trí 8" )
      Contact( "DB_Vị_trí_xe"."vị trí 5" )
      Contact( "DB_Vị_trí_xe"."vị trí 6" )
      Contact( "DB_Vị_trí_xe"."vị trí 7" )
      Coil( "DB_đầy".Tầng2 )
   END_RUNG
   // the same network as SCL:
   "DB_đầy".Tầng1 := "DB_Vị_trí_xe"."vị trí 4" AND "DB_Vị_trí_xe"."vị trí 1" AND "DB_Vị_trí_xe"."vị trí 2" AND "DB_Vị_trí_xe"."vị trí 3";
   "DB_đầy".Tầng2 := "DB_Vị_trí_xe"."vị trí 8" AND "DB_Vị_trí_xe"."vị trí 5" AND "DB_Vị_trí_xe"."vị trí 6" AND "DB_Vị_trí_xe"."vị trí 7";
END_REGION
END_FUNCTION

FUNCTION "FC_Tìm_vị_trí_tầng2" : Void   // FC6, LAD
{ S7_Optimized_Access := 'TRUE' }
VERSION : 0.1
   VAR_TEMP   // added for the SCL form of the ladder/FBD networks
      _w1 : Bool;
      _w2 : Bool;
   END_VAR
BEGIN

REGION Network 1
   // 5
